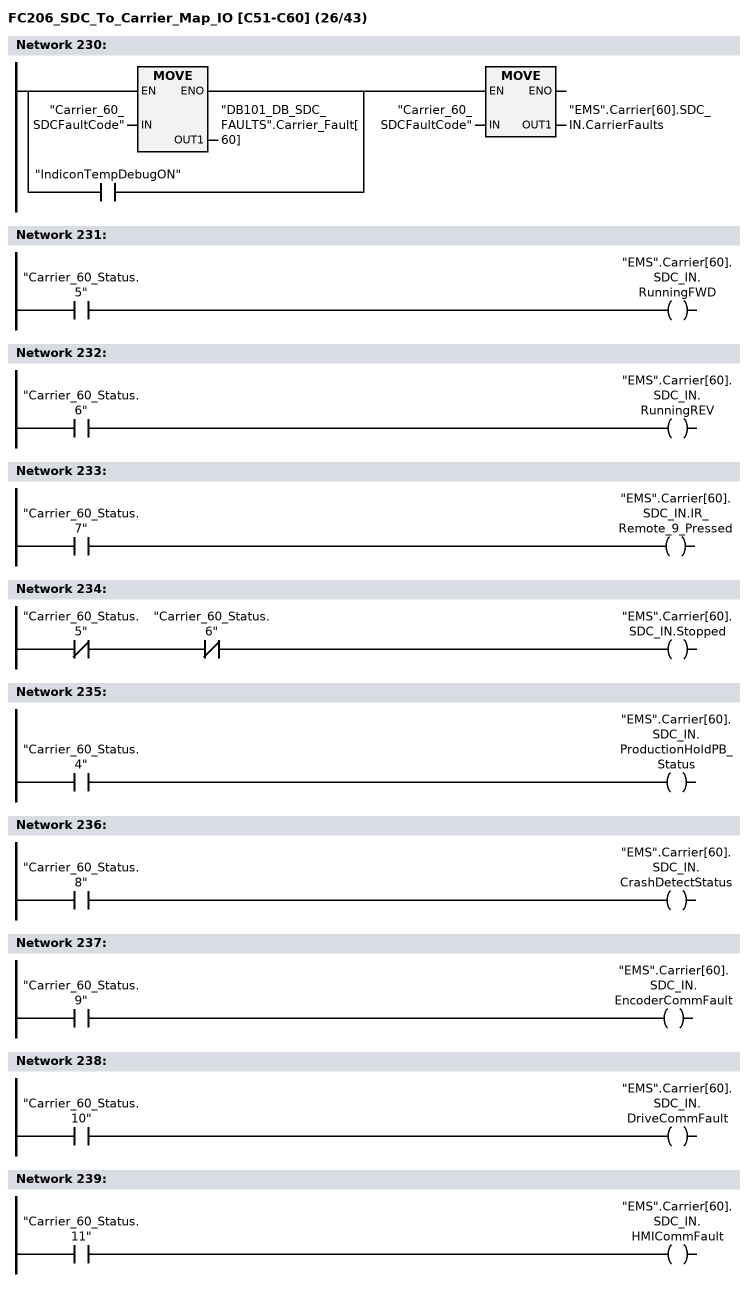
   RUNG wire#powerrail
      Move(in := "Carrier_60_SDCFaultCode", out1 => "DB101_DB_SDC_FAULTS".Carrier_Fault[60])
      wire#w1
      Move(in := "Carrier_60_SDCFaultCode", out1 => "EMS".Carrier[60].SDC_IN.CarrierFaults)
   END_RUNG
   RUNG wire#powerrail
      Contact( "IndiconTempDebugON" )
   END_RUNG wire#w1
   // the same network as SCL:
   "DB101_DB_SDC_FAULTS".Carrier_Fault[60] := "Carrier_60_SDCFaultCode";
   IF TRUE OR "IndiconTempDebugON" THEN
       "EMS".Carrier[60].SDC_IN.CarrierFaults := "Carrier_60_SDCFaultCode";
   END_IF;
END_REGION

REGION Network 231
   RUNG wire#powerrail
      Contact( "Carrier_60_Status.5" )
      Coil( "EMS".Carrier[60].SDC_IN.RunningFWD )
   END_RUNG
   // the same network as SCL:
   "EMS".Carrier[60].SDC_IN.RunningFWD := "Carrier_60_Status.5";
END_REGION

REGION Network 232
   RUNG wire#powerrail
      Contact( "Carrier_60_Status.6" )
      Coil( "EMS".Carrier[60].SDC_IN.RunningREV )
   END_RUNG
   // the same network as SCL:
   "EMS".Carrier[60].SDC_IN.RunningREV := "Carrier_60_Status.6";
END_REGION

REGION Network 233
   RUNG wire#powerrail
      Contact( "Carrier_60_Status.7" )
      Coil( "EMS".Carrier[60].SDC_IN.IR_Remote_9_Pressed )
   END_RUNG
   // the same network as SCL:
   "EMS".Carrier[60].SDC_IN.IR_Remote_9_Pressed := "Carrier_60_Status.7";
END_REGION

REGION Network 234
   RUNG wire#powerrail
      I_Contact( "Carrier_60_Status.5" )
      I_Contact( "Carrier_60_Status.6" )
      Coil( "EMS".Carrier[60].SDC_IN.Stopped )
   END_RUNG
   // the same network as SCL:
   "EMS".Carrier[60].SDC_IN.Stopped := NOT "Carrier_60_Status.5" AND NOT "Carrier_60_Status.6";
END_REGION

REGION Network 235
   RUNG wire#powerrail
      Contact( "Carrier_60_Status.4" )
      Coil( "EMS".Carrier[60].SDC_IN.ProductionHoldPB_Status )
   END_RUNG
   // the same network as SCL:
   "EMS".Carrier[60].SDC_IN.ProductionHoldPB_Status := "Carrier_60_Status.4";
END_REGION

REGION Network 236
   RUNG wire#powerrail
      Contact( "Carrier_60_Status.8" )
      Coil( "EMS".Carrier[60].SDC_IN.CrashDetectStatus )
   END_RUNG
   // the same network as SCL:
   "EMS".Carrier[60].SDC_IN.CrashDetectStatus := "Carrier_60_Status.8";
END_REGION

REGION Network 237
   RUNG wire#powerrail
      Contact( "Carrier_60_Status.9" )
      Coil( "EMS".Carrier[60].SDC_IN.EncoderCommFault )
   END_RUNG
   // the same network as SCL:
   "EMS".Carrier[60].SDC_IN.EncoderCommFault := "Carrier_60_Status.9";
END_REGION

REGION Network 238
   RUNG wire#powerrail
      Contact( "Carrier_60_Status.10" )
      Coil( "EMS".Carrier[60].SDC_IN.DriveCommFault )
   END_RUNG
   // the same network as SCL:
   "EMS".Carrier[60].SDC_IN.DriveCommFault := "Carrier_60_Status.10";
END_REGION

REGION Network 239
   RUNG wire#powerrail
      Contact( "Carrier_60_Status.11" )
      Coil( "EMS".Carrier[60].SDC_IN.HMICommFault )
   END_RUNG
   // the same network as SCL:
   "EMS".Carrier[60].SDC_IN.HMICommFault := "Carrier_60_Status.11";
END_REGION

REGION Network 240
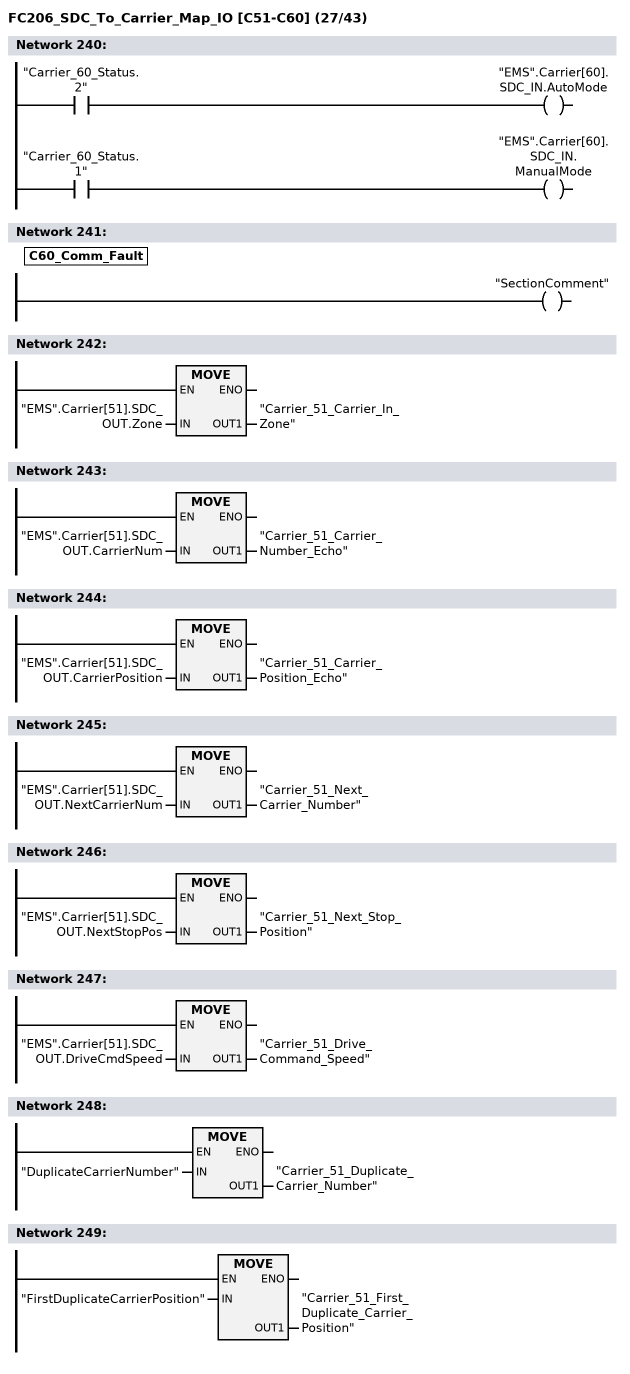
   RUNG wire#powerrail
      Contact( "Carrier_60_Status.2" )
      Coil( "EMS".Carrier[60].SDC_IN.AutoMode )
   END_RUNG
   RUNG wire#powerrail
      Contact( "Carrier_60_Status.1" )
      Coil( "EMS".Carrier[60].SDC_IN.ManualMode )
   END_RUNG
   // the same network as SCL:
   "EMS".Carrier[60].SDC_IN.AutoMode := "Carrier_60_Status.2";
   "EMS".Carrier[60].SDC_IN.ManualMode := "Carrier_60_Status.1";
END_REGION

REGION Network 241
   Label( C60_Comm_Fault )
   RUNG wire#powerrail
      Coil( "SectionComment" )
   END_RUNG
   // the same network as SCL:
   C60_Comm_Fault:
   "SectionComment" := TRUE;
END_REGION

REGION Network 242
   RUNG wire#powerrail
      Move(in := "EMS".Carrier[51].SDC_OUT.Zone, out1 => "Carrier_51_Carrier_In_Zone")
   END_RUNG
   // the same network as SCL:
   "Carrier_51_Carrier_In_Zone" := "EMS".Carrier[51].SDC_OUT.Zone;
END_REGION

REGION Network 243
   RUNG wire#powerrail
      Move(in := "EMS".Carrier[51].SDC_OUT.CarrierNum, out1 => "Carrier_51_Carrier_Number_Echo")
   END_RUNG
   // the same network as SCL:
   "Carrier_51_Carrier_Number_Echo" := "EMS".Carrier[51].SDC_OUT.CarrierNum;
END_REGION

REGION Network 244
   RUNG wire#powerrail
      Move(in := "EMS".Carrier[51].SDC_OUT.CarrierPosition, out1 => "Carrier_51_Carrier_Position_Echo")
   END_RUNG
   // the same network as SCL:
   "Carrier_51_Carrier_Position_Echo" := "EMS".Carrier[51].SDC_OUT.CarrierPosition;
END_REGION

REGION Network 245
   RUNG wire#powerrail
      Move(in := "EMS".Carrier[51].SDC_OUT.NextCarrierNum, out1 => "Carrier_51_Next_Carrier_Number")
   END_RUNG
   // the same network as SCL:
   "Carrier_51_Next_Carrier_Number" := "EMS".Carrier[51].SDC_OUT.NextCarrierNum;
END_REGION

REGION Network 246
   RUNG wire#powerrail
      Move(in := "EMS".Carrier[51].SDC_OUT.NextStopPos, out1 => "Carrier_51_Next_Stop_Position")
   END_RUNG
   // the same network as SCL:
   "Carrier_51_Next_Stop_Position" := "EMS".Carrier[51].SDC_OUT.NextStopPos;
END_REGION

REGION Network 247
   RUNG wire#powerrail
      Move(in := "EMS".Carrier[51].SDC_OUT.DriveCmdSpeed, out1 => "Carrier_51_Drive_Command_Speed")
   END_RUNG
   // the same network as SCL:
   "Carrier_51_Drive_Command_Speed" := "EMS".Carrier[51].SDC_OUT.DriveCmdSpeed;
END_REGION

REGION Network 248
   RUNG wire#powerrail
      Move(in := "DuplicateCarrierNumber", out1 => "Carrier_51_Duplicate_Carrier_Number")
   END_RUNG
   // the same network as SCL:
   "Carrier_51_Duplicate_Carrier_Number" := "DuplicateCarrierNumber";
END_REGION

REGION Network 249
   RUNG wire#powerrail
      Move(in := "FirstDuplicateCarrierPosition", out1 => "Carrier_51_First_Duplicate_Carrier_Position")
   END_RUNG
   // the same network as SCL:
   "Carrier_51_First_Duplicate_Carrier_Position" := "FirstDuplicateCarrierPosition";
END_REGION

REGION Network 250
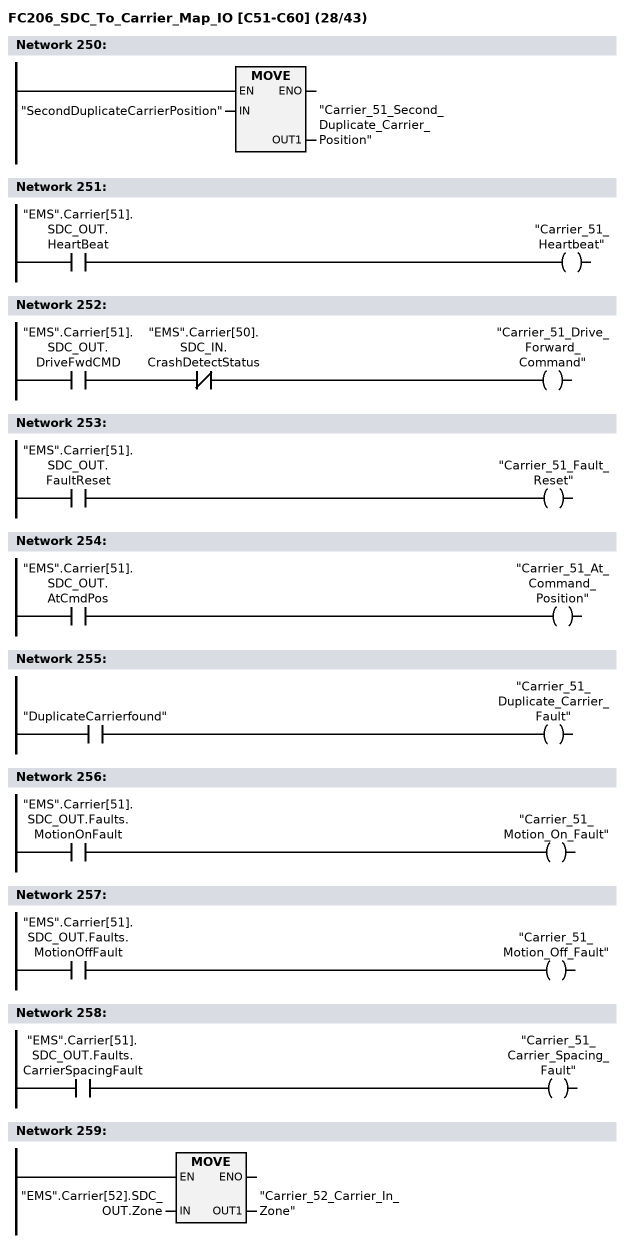
   RUNG wire#powerrail
      Move(in := "SecondDuplicateCarrierPosition", out1 => "Carrier_51_Second_Duplicate_Carrier_Position")
   END_RUNG
   // the same network as SCL:
   "Carrier_51_Second_Duplicate_Carrier_Position" := "SecondDuplicateCarrierPosition";
END_REGION

REGION Network 251
   RUNG wire#powerrail
      Contact( "EMS".Carrier[51].SDC_OUT.HeartBeat )
      Coil( "Carrier_51_Heartbeat" )
   END_RUNG
   // the same network as SCL:
   "Carrier_51_Heartbeat" := "EMS".Carrier[51].SDC_OUT.HeartBeat;
END_REGION

REGION Network 252
   RUNG wire#powerrail
      Contact( "EMS".Carrier[51].SDC_OUT.DriveFwdCMD )
      I_Contact( "EMS".Carrier[50].SDC_IN.CrashDetectStatus )
      Coil( "Carrier_51_Drive_Forward_Command" )
   END_RUNG
   // the same network as SCL:
   "Carrier_51_Drive_Forward_Command" := "EMS".Carrier[51].SDC_OUT.DriveFwdCMD AND NOT "EMS".Carrier[50].SDC_IN.CrashDetectStatus;
END_REGION

REGION Network 253
   RUNG wire#powerrail
      Contact( "EMS".Carrier[51].SDC_OUT.FaultReset )
      Coil( "Carrier_51_Fault_Reset" )
   END_RUNG
   // the same network as SCL:
   "Carrier_51_Fault_Reset" := "EMS".Carrier[51].SDC_OUT.FaultReset;
END_REGION

REGION Network 254
   RUNG wire#powerrail
      Contact( "EMS".Carrier[51].SDC_OUT.AtCmdPos )
      Coil( "Carrier_51_At_Command_Position" )
   END_RUNG
   // the same network as SCL:
   "Carrier_51_At_Command_Position" := "EMS".Carrier[51].SDC_OUT.AtCmdPos;
END_REGION

REGION Network 255
   RUNG wire#powerrail
      Contact( "DuplicateCarrierfound" )
      Coil( "Carrier_51_Duplicate_Carrier_Fault" )
   END_RUNG
   // the same network as SCL:
   "Carrier_51_Duplicate_Carrier_Fault" := "DuplicateCarrierfound";
END_REGION

REGION Network 256
   RUNG wire#powerrail
      Contact( "EMS".Carrier[51].SDC_OUT.Faults.MotionOnFault )
      Coil( "Carrier_51_Motion_On_Fault" )
   END_RUNG
   // the same network as SCL:
   "Carrier_51_Motion_On_Fault" := "EMS".Carrier[51].SDC_OUT.Faults.MotionOnFault;
END_REGION

REGION Network 257
   RUNG wire#powerrail
      Contact( "EMS".Carrier[51].SDC_OUT.Faults.MotionOffFault )
      Coil( "Carrier_51_Motion_Off_Fault" )
   END_RUNG
   // the same network as SCL:
   "Carrier_51_Motion_Off_Fault" := "EMS".Carrier[51].SDC_OUT.Faults.MotionOffFault;
END_REGION

REGION Network 258
   RUNG wire#powerrail
      Contact( "EMS".Carrier[51].SDC_OUT.Faults.CarrierSpacingFault )
      Coil( "Carrier_51_Carrier_Spacing_Fault" )
   END_RUNG
   // the same network as SCL:
   "Carrier_51_Carrier_Spacing_Fault" := "EMS".Carrier[51].SDC_OUT.Faults.CarrierSpacingFault;
END_REGION

REGION Network 259
   RUNG wire#powerrail
      Move(in := "EMS".Carrier[52].SDC_OUT.Zone, out1 => "Carrier_52_Carrier_In_Zone")
   END_RUNG
   // the same network as SCL:
   "Carrier_52_Carrier_In_Zone" := "EMS".Carrier[52].SDC_OUT.Zone;
END_REGION

REGION Network 260
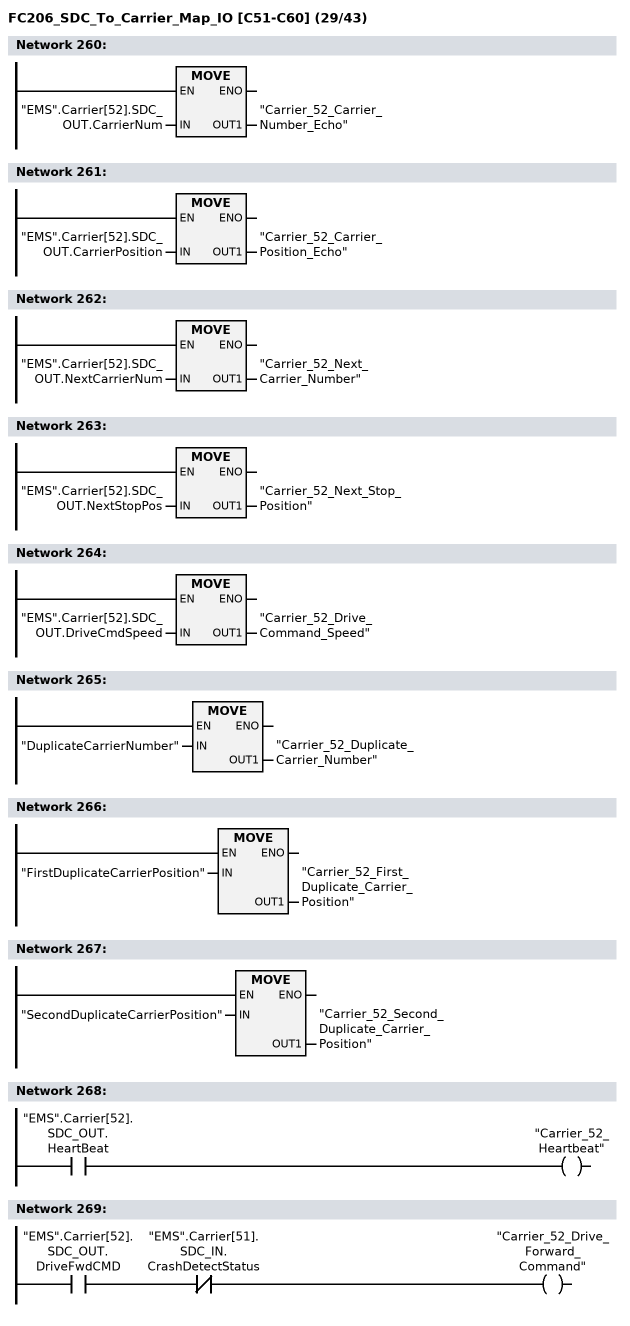
   RUNG wire#powerrail
      Move(in := "EMS".Carrier[52].SDC_OUT.CarrierNum, out1 => "Carrier_52_Carrier_Number_Echo")
   END_RUNG
   // the same network as SCL:
   "Carrier_52_Carrier_Number_Echo" := "EMS".Carrier[52].SDC_OUT.CarrierNum;
END_REGION

REGION Network 261
   RUNG wire#powerrail
      Move(in := "EMS".Carrier[52].SDC_OUT.CarrierPosition, out1 => "Carrier_52_Carrier_Position_Echo")
   END_RUNG
   // the same network as SCL:
   "Carrier_52_Carrier_Position_Echo" := "EMS".Carrier[52].SDC_OUT.CarrierPosition;
END_REGION

REGION Network 262
   RUNG wire#powerrail
      Move(in := "EMS".Carrier[52].SDC_OUT.NextCarrierNum, out1 => "Carrier_52_Next_Carrier_Number")
   END_RUNG
   // the same network as SCL:
   "Carrier_52_Next_Carrier_Number" := "EMS".Carrier[52].SDC_OUT.NextCarrierNum;
END_REGION

REGION Network 263
   RUNG wire#powerrail
      Move(in := "EMS".Carrier[52].SDC_OUT.NextStopPos, out1 => "Carrier_52_Next_Stop_Position")
   END_RUNG
   // the same network as SCL:
   "Carrier_52_Next_Stop_Position" := "EMS".Carrier[52].SDC_OUT.NextStopPos;
END_REGION

REGION Network 264
   RUNG wire#powerrail
      Move(in := "EMS".Carrier[52].SDC_OUT.DriveCmdSpeed, out1 => "Carrier_52_Drive_Command_Speed")
   END_RUNG
   // the same network as SCL:
   "Carrier_52_Drive_Command_Speed" := "EMS".Carrier[52].SDC_OUT.DriveCmdSpeed;
END_REGION

REGION Network 265
   RUNG wire#powerrail
      Move(in := "DuplicateCarrierNumber", out1 => "Carrier_52_Duplicate_Carrier_Number")
   END_RUNG
   // the same network as SCL:
   "Carrier_52_Duplicate_Carrier_Number" := "DuplicateCarrierNumber";
END_REGION

REGION Network 266
   RUNG wire#powerrail
      Move(in := "FirstDuplicateCarrierPosition", out1 => "Carrier_52_First_Duplicate_Carrier_Position")
   END_RUNG
   // the same network as SCL:
   "Carrier_52_First_Duplicate_Carrier_Position" := "FirstDuplicateCarrierPosition";
END_REGION

REGION Network 267
   RUNG wire#powerrail
      Move(in := "SecondDuplicateCarrierPosition", out1 => "Carrier_52_Second_Duplicate_Carrier_Position")
   END_RUNG
   // the same network as SCL:
   "Carrier_52_Second_Duplicate_Carrier_Position" := "SecondDuplicateCarrierPosition";
END_REGION

REGION Network 268
   RUNG wire#powerrail
      Contact( "EMS".Carrier[52].SDC_OUT.HeartBeat )
      Coil( "Carrier_52_Heartbeat" )
   END_RUNG
   // the same network as SCL:
   "Carrier_52_Heartbeat" := "EMS".Carrier[52].SDC_OUT.HeartBeat;
END_REGION

REGION Network 269
   RUNG wire#powerrail
      Contact( "EMS".Carrier[52].SDC_OUT.DriveFwdCMD )
      I_Contact( "EMS".Carrier[51].SDC_IN.CrashDetectStatus )
      Coil( "Carrier_52_Drive_Forward_Command" )
   END_RUNG
   // the same network as SCL:
   "Carrier_52_Drive_Forward_Command" := "EMS".Carrier[52].SDC_OUT.DriveFwdCMD AND NOT "EMS".Carrier[51].SDC_IN.CrashDetectStatus;
END_REGION

REGION Network 270
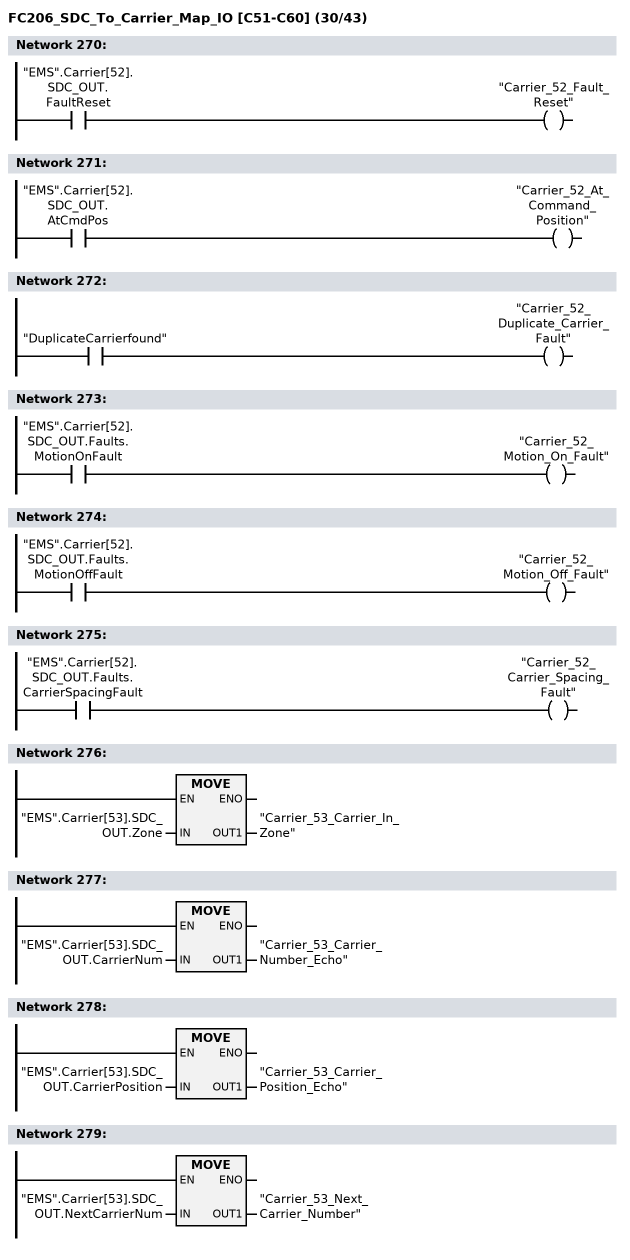
   RUNG wire#powerrail
      Contact( "EMS".Carrier[52].SDC_OUT.FaultReset )
      Coil( "Carrier_52_Fault_Reset" )
   END_RUNG
   // the same network as SCL:
   "Carrier_52_Fault_Reset" := "EMS".Carrier[52].SDC_OUT.FaultReset;
END_REGION

REGION Network 271
   RUNG wire#powerrail
      Contact( "EMS".Carrier[52].SDC_OUT.AtCmdPos )
      Coil( "Carrier_52_At_Command_Position" )
   END_RUNG
   // the same network as SCL:
   "Carrier_52_At_Command_Position" := "EMS".Carrier[52].SDC_OUT.AtCmdPos;
END_REGION

REGION Network 272
   RUNG wire#powerrail
      Contact( "DuplicateCarrierfound" )
      Coil( "Carrier_52_Duplicate_Carrier_Fault" )
   END_RUNG
   // the same network as SCL:
   "Carrier_52_Duplicate_Carrier_Fault" := "DuplicateCarrierfound";
END_REGION

REGION Network 273
   RUNG wire#powerrail
      Contact( "EMS".Carrier[52].SDC_OUT.Faults.MotionOnFault )
      Coil( "Carrier_52_Motion_On_Fault" )
   END_RUNG
   // the same network as SCL:
   "Carrier_52_Motion_On_Fault" := "EMS".Carrier[52].SDC_OUT.Faults.MotionOnFault;
END_REGION

REGION Network 274
   RUNG wire#powerrail
      Contact( "EMS".Carrier[52].SDC_OUT.Faults.MotionOffFault )
      Coil( "Carrier_52_Motion_Off_Fault" )
   END_RUNG
   // the same network as SCL:
   "Carrier_52_Motion_Off_Fault" := "EMS".Carrier[52].SDC_OUT.Faults.MotionOffFault;
END_REGION

REGION Network 275
   RUNG wire#powerrail
      Contact( "EMS".Carrier[52].SDC_OUT.Faults.CarrierSpacingFault )
      Coil( "Carrier_52_Carrier_Spacing_Fault" )
   END_RUNG
   // the same network as SCL:
   "Carrier_52_Carrier_Spacing_Fault" := "EMS".Carrier[52].SDC_OUT.Faults.CarrierSpacingFault;
END_REGION

REGION Network 276
   RUNG wire#powerrail
      Move(in := "EMS".Carrier[53].SDC_OUT.Zone, out1 => "Carrier_53_Carrier_In_Zone")
   END_RUNG
   // the same network as SCL:
   "Carrier_53_Carrier_In_Zone" := "EMS".Carrier[53].SDC_OUT.Zone;
END_REGION

REGION Network 277
   RUNG wire#powerrail
      Move(in := "EMS".Carrier[53].SDC_OUT.CarrierNum, out1 => "Carrier_53_Carrier_Number_Echo")
   END_RUNG
   // the same network as SCL:
   "Carrier_53_Carrier_Number_Echo" := "EMS".Carrier[53].SDC_OUT.CarrierNum;
END_REGION

REGION Network 278
   RUNG wire#powerrail
      Move(in := "EMS".Carrier[53].SDC_OUT.CarrierPosition, out1 => "Carrier_53_Carrier_Position_Echo")
   END_RUNG
   // the same network as SCL:
   "Carrier_53_Carrier_Position_Echo" := "EMS".Carrier[53].SDC_OUT.CarrierPosition;
END_REGION

REGION Network 279
   RUNG wire#powerrail
      Move(in := "EMS".Carrier[53].SDC_OUT.NextCarrierNum, out1 => "Carrier_53_Next_Carrier_Number")
   END_RUNG
   // the same network as SCL:
   "Carrier_53_Next_Carrier_Number" := "EMS".Carrier[53].SDC_OUT.NextCarrierNum;
END_REGION

REGION Network 280
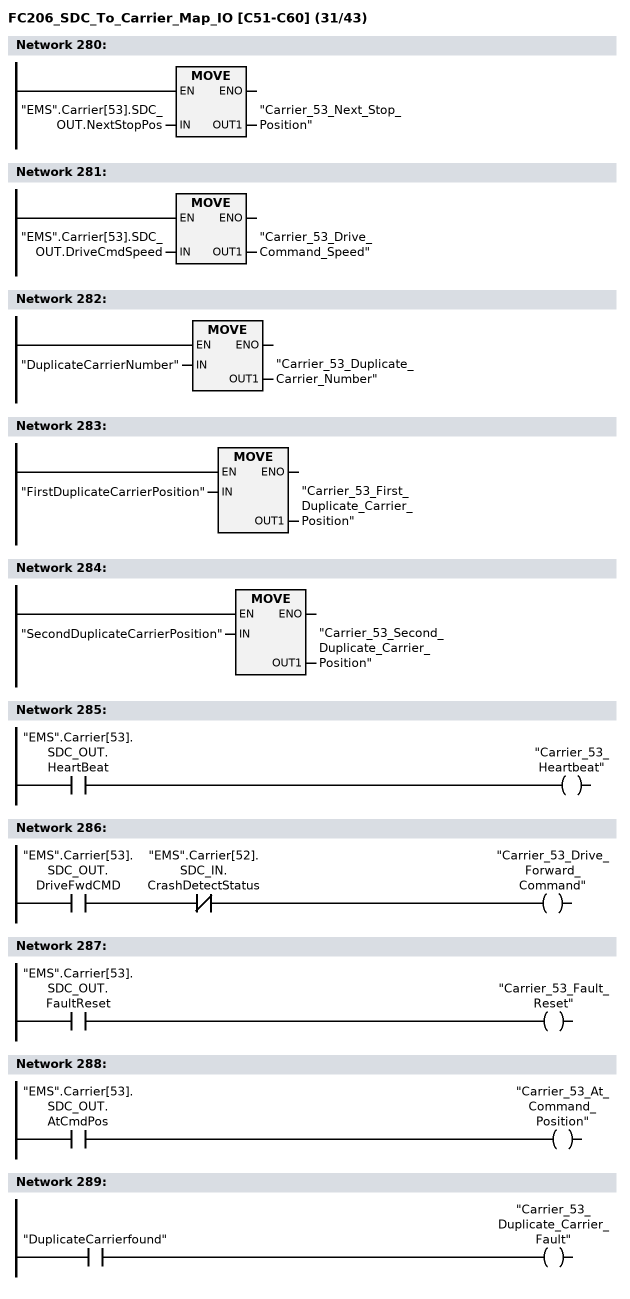
   RUNG wire#powerrail
      Move(in := "EMS".Carrier[53].SDC_OUT.NextStopPos, out1 => "Carrier_53_Next_Stop_Position")
   END_RUNG
   // the same network as SCL:
   "Carrier_53_Next_Stop_Position" := "EMS".Carrier[53].SDC_OUT.NextStopPos;
END_REGION

REGION Network 281
   RUNG wire#powerrail
      Move(in := "EMS".Carrier[53].SDC_OUT.DriveCmdSpeed, out1 => "Carrier_53_Drive_Command_Speed")
   END_RUNG
   // the same network as SCL:
   "Carrier_53_Drive_Command_Speed" := "EMS".Carrier[53].SDC_OUT.DriveCmdSpeed;
END_REGION

REGION Network 282
   RUNG wire#powerrail
      Move(in := "DuplicateCarrierNumber", out1 => "Carrier_53_Duplicate_Carrier_Number")
   END_RUNG
   // the same network as SCL:
   "Carrier_53_Duplicate_Carrier_Number" := "DuplicateCarrierNumber";
END_REGION

REGION Network 283
   RUNG wire#powerrail
      Move(in := "FirstDuplicateCarrierPosition", out1 => "Carrier_53_First_Duplicate_Carrier_Position")
   END_RUNG
   // the same network as SCL:
   "Carrier_53_First_Duplicate_Carrier_Position" := "FirstDuplicateCarrierPosition";
END_REGION

REGION Network 284
   RUNG wire#powerrail
      Move(in := "SecondDuplicateCarrierPosition", out1 => "Carrier_53_Second_Duplicate_Carrier_Position")
   END_RUNG
   // the same network as SCL:
   "Carrier_53_Second_Duplicate_Carrier_Position" := "SecondDuplicateCarrierPosition";
END_REGION

REGION Network 285
   RUNG wire#powerrail
      Contact( "EMS".Carrier[53].SDC_OUT.HeartBeat )
      Coil( "Carrier_53_Heartbeat" )
   END_RUNG
   // the same network as SCL:
   "Carrier_53_Heartbeat" := "EMS".Carrier[53].SDC_OUT.HeartBeat;
END_REGION

REGION Network 286
   RUNG wire#powerrail
      Contact( "EMS".Carrier[53].SDC_OUT.DriveFwdCMD )
      I_Contact( "EMS".Carrier[52].SDC_IN.CrashDetectStatus )
      Coil( "Carrier_53_Drive_Forward_Command" )
   END_RUNG
   // the same network as SCL:
   "Carrier_53_Drive_Forward_Command" := "EMS".Carrier[53].SDC_OUT.DriveFwdCMD AND NOT "EMS".Carrier[52].SDC_IN.CrashDetectStatus;
END_REGION

REGION Network 287
   RUNG wire#powerrail
      Contact( "EMS".Carrier[53].SDC_OUT.FaultReset )
      Coil( "Carrier_53_Fault_Reset" )
   END_RUNG
   // the same network as SCL:
   "Carrier_53_Fault_Reset" := "EMS".Carrier[53].SDC_OUT.FaultReset;
END_REGION

REGION Network 288
   RUNG wire#powerrail
      Contact( "EMS".Carrier[53].SDC_OUT.AtCmdPos )
      Coil( "Carrier_53_At_Command_Position" )
   END_RUNG
   // the same network as SCL:
   "Carrier_53_At_Command_Position" := "EMS".Carrier[53].SDC_OUT.AtCmdPos;
END_REGION

REGION Network 289
   RUNG wire#powerrail
      Contact( "DuplicateCarrierfound" )
      Coil( "Carrier_53_Duplicate_Carrier_Fault" )
   END_RUNG
   // the same network as SCL:
   "Carrier_53_Duplicate_Carrier_Fault" := "DuplicateCarrierfound";
END_REGION

REGION Network 290
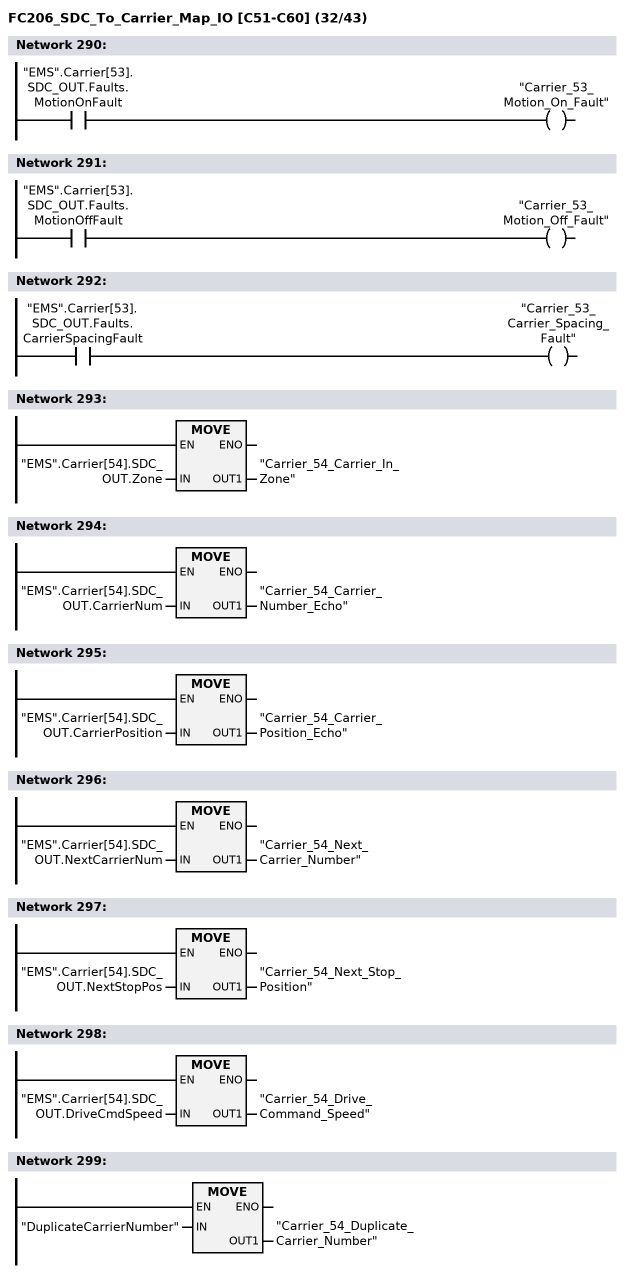
   RUNG wire#powerrail
      Contact( "EMS".Carrier[53].SDC_OUT.Faults.MotionOnFault )
      Coil( "Carrier_53_Motion_On_Fault" )
   END_RUNG
   // the same network as SCL:
   "Carrier_53_Motion_On_Fault" := "EMS".Carrier[53].SDC_OUT.Faults.MotionOnFault;
END_REGION

REGION Network 291
   RUNG wire#powerrail
      Contact( "EMS".Carrier[53].SDC_OUT.Faults.MotionOffFault )
      Coil( "Carrier_53_Motion_Off_Fault" )
   END_RUNG
   // the same network as SCL:
   "Carrier_53_Motion_Off_Fault" := "EMS".Carrier[53].SDC_OUT.Faults.MotionOffFault;
END_REGION

REGION Network 292
   RUNG wire#powerrail
      Contact( "EMS".Carrier[53].SDC_OUT.Faults.CarrierSpacingFault )
      Coil( "Carrier_53_Carrier_Spacing_Fault" )
   END_RUNG
   // the same network as SCL:
   "Carrier_53_Carrier_Spacing_Fault" := "EMS".Carrier[53].SDC_OUT.Faults.CarrierSpacingFault;
END_REGION

REGION Network 293
   RUNG wire#powerrail
      Move(in := "EMS".Carrier[54].SDC_OUT.Zone, out1 => "Carrier_54_Carrier_In_Zone")
   END_RUNG
   // the same network as SCL:
   "Carrier_54_Carrier_In_Zone" := "EMS".Carrier[54].SDC_OUT.Zone;
END_REGION

REGION Network 294
   RUNG wire#powerrail
      Move(in := "EMS".Carrier[54].SDC_OUT.CarrierNum, out1 => "Carrier_54_Carrier_Number_Echo")
   END_RUNG
   // the same network as SCL:
   "Carrier_54_Carrier_Number_Echo" := "EMS".Carrier[54].SDC_OUT.CarrierNum;
END_REGION

REGION Network 295
   RUNG wire#powerrail
      Move(in := "EMS".Carrier[54].SDC_OUT.CarrierPosition, out1 => "Carrier_54_Carrier_Position_Echo")
   END_RUNG
   // the same network as SCL:
   "Carrier_54_Carrier_Position_Echo" := "EMS".Carrier[54].SDC_OUT.CarrierPosition;
END_REGION

REGION Network 296
   RUNG wire#powerrail
      Move(in := "EMS".Carrier[54].SDC_OUT.NextCarrierNum, out1 => "Carrier_54_Next_Carrier_Number")
   END_RUNG
   // the same network as SCL:
   "Carrier_54_Next_Carrier_Number" := "EMS".Carrier[54].SDC_OUT.NextCarrierNum;
END_REGION

REGION Network 297
   RUNG wire#powerrail
      Move(in := "EMS".Carrier[54].SDC_OUT.NextStopPos, out1 => "Carrier_54_Next_Stop_Position")
   END_RUNG
   // the same network as SCL:
   "Carrier_54_Next_Stop_Position" := "EMS".Carrier[54].SDC_OUT.NextStopPos;
END_REGION

REGION Network 298
   RUNG wire#powerrail
      Move(in := "EMS".Carrier[54].SDC_OUT.DriveCmdSpeed, out1 => "Carrier_54_Drive_Command_Speed")
   END_RUNG
   // the same network as SCL:
   "Carrier_54_Drive_Command_Speed" := "EMS".Carrier[54].SDC_OUT.DriveCmdSpeed;
END_REGION

REGION Network 299
   RUNG wire#powerrail
      Move(in := "DuplicateCarrierNumber", out1 => "Carrier_54_Duplicate_Carrier_Number")
   END_RUNG
   // the same network as SCL:
   "Carrier_54_Duplicate_Carrier_Number" := "DuplicateCarrierNumber";
END_REGION

REGION Network 300
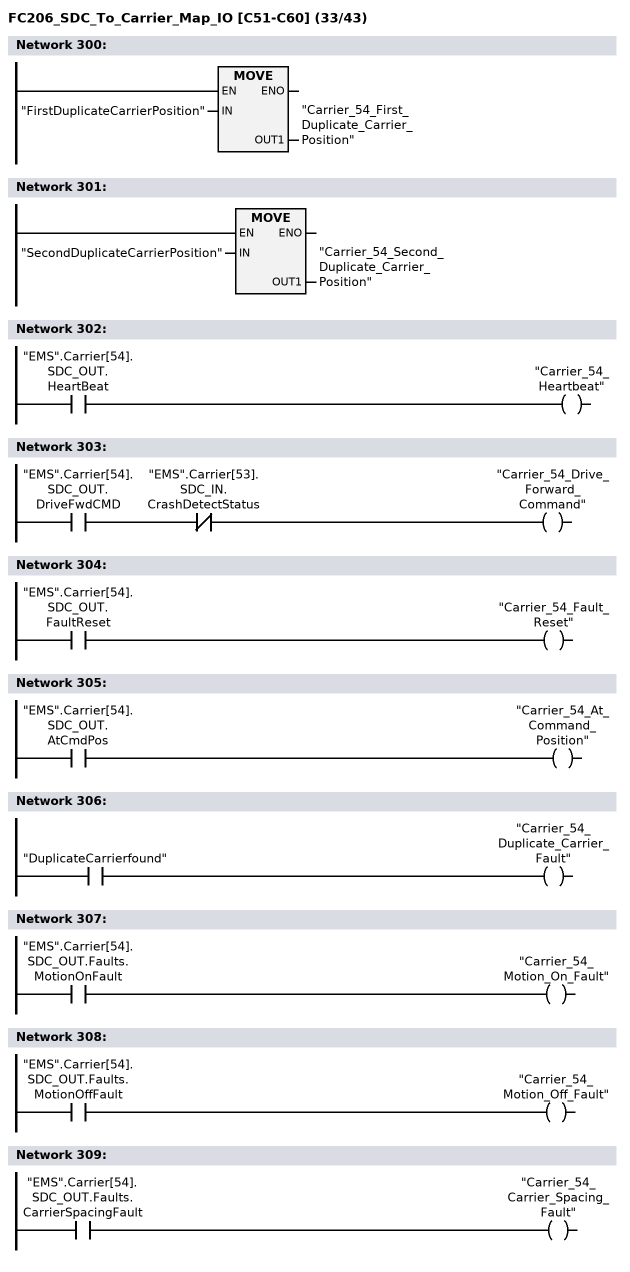
   RUNG wire#powerrail
      Move(in := "FirstDuplicateCarrierPosition", out1 => "Carrier_54_First_Duplicate_Carrier_Position")
   END_RUNG
   // the same network as SCL:
   "Carrier_54_First_Duplicate_Carrier_Position" := "FirstDuplicateCarrierPosition";
END_REGION

REGION Network 301
   RUNG wire#powerrail
      Move(in := "SecondDuplicateCarrierPosition", out1 => "Carrier_54_Second_Duplicate_Carrier_Position")
   END_RUNG
   // the same network as SCL:
   "Carrier_54_Second_Duplicate_Carrier_Position" := "SecondDuplicateCarrierPosition";
END_REGION

REGION Network 302
   RUNG wire#powerrail
      Contact( "EMS".Carrier[54].SDC_OUT.HeartBeat )
      Coil( "Carrier_54_Heartbeat" )
   END_RUNG
   // the same network as SCL:
   "Carrier_54_Heartbeat" := "EMS".Carrier[54].SDC_OUT.HeartBeat;
END_REGION

REGION Network 303
   RUNG wire#powerrail
      Contact( "EMS".Carrier[54].SDC_OUT.DriveFwdCMD )
      I_Contact( "EMS".Carrier[53].SDC_IN.CrashDetectStatus )
      Coil( "Carrier_54_Drive_Forward_Command" )
   END_RUNG
   // the same network as SCL:
   "Carrier_54_Drive_Forward_Command" := "EMS".Carrier[54].SDC_OUT.DriveFwdCMD AND NOT "EMS".Carrier[53].SDC_IN.CrashDetectStatus;
END_REGION

REGION Network 304
   RUNG wire#powerrail
      Contact( "EMS".Carrier[54].SDC_OUT.FaultReset )
      Coil( "Carrier_54_Fault_Reset" )
   END_RUNG
   // the same network as SCL:
   "Carrier_54_Fault_Reset" := "EMS".Carrier[54].SDC_OUT.FaultReset;
END_REGION

REGION Network 305
   RUNG wire#powerrail
      Contact( "EMS".Carrier[54].SDC_OUT.AtCmdPos )
      Coil( "Carrier_54_At_Command_Position" )
   END_RUNG
   // the same network as SCL:
   "Carrier_54_At_Command_Position" := "EMS".Carrier[54].SDC_OUT.AtCmdPos;
END_REGION

REGION Network 306
   RUNG wire#powerrail
      Contact( "DuplicateCarrierfound" )
      Coil( "Carrier_54_Duplicate_Carrier_Fault" )
   END_RUNG
   // the same network as SCL:
   "Carrier_54_Duplicate_Carrier_Fault" := "DuplicateCarrierfound";
END_REGION

REGION Network 307
   RUNG wire#powerrail
      Contact( "EMS".Carrier[54].SDC_OUT.Faults.MotionOnFault )
      Coil( "Carrier_54_Motion_On_Fault" )
   END_RUNG
   // the same network as SCL:
   "Carrier_54_Motion_On_Fault" := "EMS".Carrier[54].SDC_OUT.Faults.MotionOnFault;
END_REGION

REGION Network 308
   RUNG wire#powerrail
      Contact( "EMS".Carrier[54].SDC_OUT.Faults.MotionOffFault )
      Coil( "Carrier_54_Motion_Off_Fault" )
   END_RUNG
   // the same network as SCL:
   "Carrier_54_Motion_Off_Fault" := "EMS".Carrier[54].SDC_OUT.Faults.MotionOffFault;
END_REGION

REGION Network 309
   RUNG wire#powerrail
      Contact( "EMS".Carrier[54].SDC_OUT.Faults.CarrierSpacingFault )
      Coil( "Carrier_54_Carrier_Spacing_Fault" )
   END_RUNG
   // the same network as SCL:
   "Carrier_54_Carrier_Spacing_Fault" := "EMS".Carrier[54].SDC_OUT.Faults.CarrierSpacingFault;
END_REGION

REGION Network 310